   "FB_Z200Conveyor_M211_iDB"(IN_xCycleON := "Z201".ST_xCycleON,
                              IN_xCycleONDel := "Z201".ST_xCycleONDelayed,
                              IN_xFaultsEnabled := "Z201".ST_xFaultsEnabled,
                              IN_xResetAlarms := "Z201".tmOFF_ResetAlarm.OUT_xDone,
                              IN_xAccelation:=FALSE,
                              IN_rgtMotorConfig := #TMP_rgtMotorConfig);
END_REGION

REGION Network 12 (SCL): Outputs Z200
   "ZUPS_Output"();
   "Z201_Output"();
   "Z200_Output"();

   "Output_Z201_Idevice"();
END_REGION
END_ORGANIZATION_BLOCK

// folder: TaskMedium

ORGANIZATION_BLOCK "OBx_TaskMedium"   // OB31, LAD, CyclicInterrupt
{ S7_Optimized_Access := 'TRUE' }
VERSION : 0.1
   VAR_INPUT
      Initial_Call : Bool;   // Initial call of this OB
      Event_Count : Int;   // Events discarded
   END_VAR
   VAR_TEMP
      TMP_iRetVal : Int;
      TMP_xDummy : Bool;
   END_VAR
BEGIN

REGION Network 1: Initialize
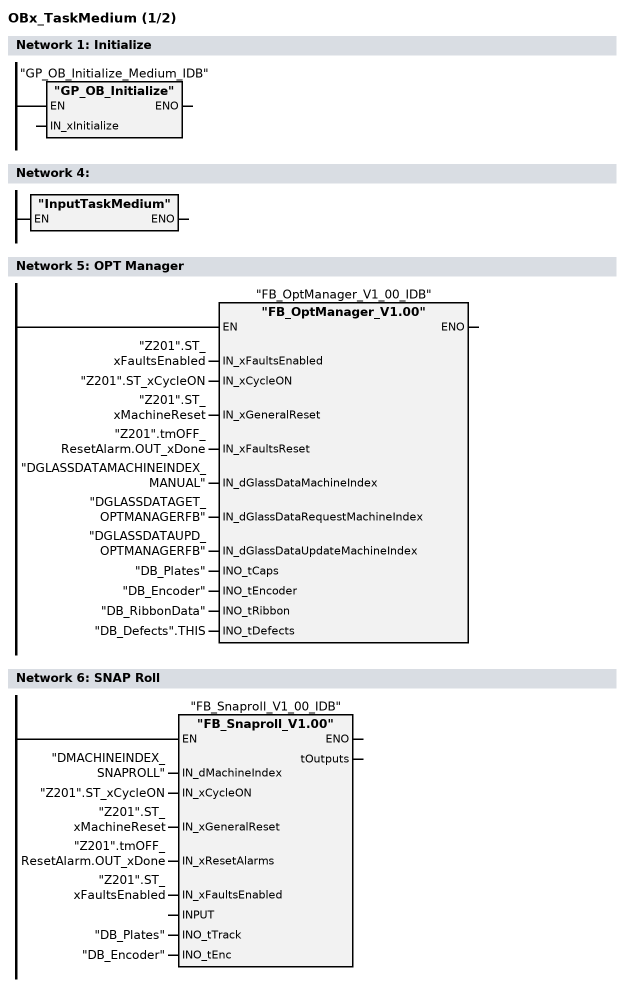
   RUNG wire#powerrail
      "GP_OB_Initialize_Medium_IDB"(IN_xInitialize :=)
   END_RUNG
   // the same network as SCL:
   "GP_OB_Initialize_Medium_IDB"();   // "GP_OB_Initialize"
END_REGION

REGION Network 2: OB Scan
END_REGION

REGION Network 3 (SCL): Message call

   "RP_OB_TaskMediumToOpt"(FALSE);
   "RP_OB_TaskMediumFromOpt"(FALSE);
END_REGION

REGION Network 4
   RUNG wire#powerrail
      "InputTaskMedium"()
   END_RUNG
   // the same network as SCL:
   "InputTaskMedium"();
END_REGION

REGION Network 5: OPT Manager
   RUNG wire#powerrail
      "FB_OptManager_V1_00_IDB"(IN_xFaultsEnabled := "Z201".ST_xFaultsEnabled, IN_xCycleON := "Z201".ST_xCycleON, IN_xGeneralReset := "Z201".ST_xMachineReset, IN_xFaultsReset := "Z201".tmOFF_ResetAlarm.OUT_xDone, IN_dGlassDataMachineIndex := "DGLASSDATAMACHINEINDEX_MANUAL", IN_dGlassDataRequestMachineIndex := "DGLASSDATAGET_OPTMANAGERFB", IN_dGlassDataUpdateMachineIndex := "DGLASSDATAUPD_OPTMANAGERFB", INO_tCaps := "DB_Plates", INO_tEncoder := "DB_Encoder", INO_tRibbon := "DB_RibbonData", INO_tDefects := "DB_Defects".THIS)
   END_RUNG
   // the same network as SCL:
   "FB_OptManager_V1_00_IDB"(IN_xFaultsEnabled := "Z201".ST_xFaultsEnabled,   // "FB_OptManager_V1.00"
                           IN_xCycleON := "Z201".ST_xCycleON,
                           IN_xGeneralReset := "Z201".ST_xMachineReset,
                           IN_xFaultsReset := "Z201".tmOFF_ResetAlarm.OUT_xDone,
                           IN_dGlassDataMachineIndex := "DGLASSDATAMACHINEINDEX_MANUAL",
                           IN_dGlassDataRequestMachineIndex := "DGLASSDATAGET_OPTMANAGERFB",
                           IN_dGlassDataUpdateMachineIndex := "DGLASSDATAUPD_OPTMANAGERFB",
                           INO_tCaps := "DB_Plates",
                           INO_tEncoder := "DB_Encoder",
                           INO_tRibbon := "DB_RibbonData",
                           INO_tDefects := "DB_Defects".THIS);
END_REGION

REGION Network 6: SNAP Roll
   RUNG wire#powerrail
      "FB_Snaproll_V1_00_IDB"(IN_dMachineIndex := "DMACHINEINDEX_SNAPROLL", IN_xCycleON := "Z201".ST_xCycleON, IN_xGeneralReset := "Z201".ST_xMachineReset, IN_xResetAlarms := "Z201".tmOFF_ResetAlarm.OUT_xDone, IN_xFaultsEnabled := "Z201".ST_xFaultsEnabled, INPUT :=, INO_tTrack := "DB_Plates", INO_tEnc := "DB_Encoder", tOutputs =>)
   END_RUNG
   // the same network as SCL:
   "FB_Snaproll_V1_00_IDB"(IN_dMachineIndex := "DMACHINEINDEX_SNAPROLL",   // "FB_Snaproll_V1.00"
                           IN_xCycleON := "Z201".ST_xCycleON,
                           IN_xGeneralReset := "Z201".ST_xMachineReset,
                           IN_xResetAlarms := "Z201".tmOFF_ResetAlarm.OUT_xDone,
                           IN_xFaultsEnabled := "Z201".ST_xFaultsEnabled,
                           INO_tTrack := "DB_Plates",
                           INO_tEnc := "DB_Encoder");
END_REGION

REGION Network 7: Z300
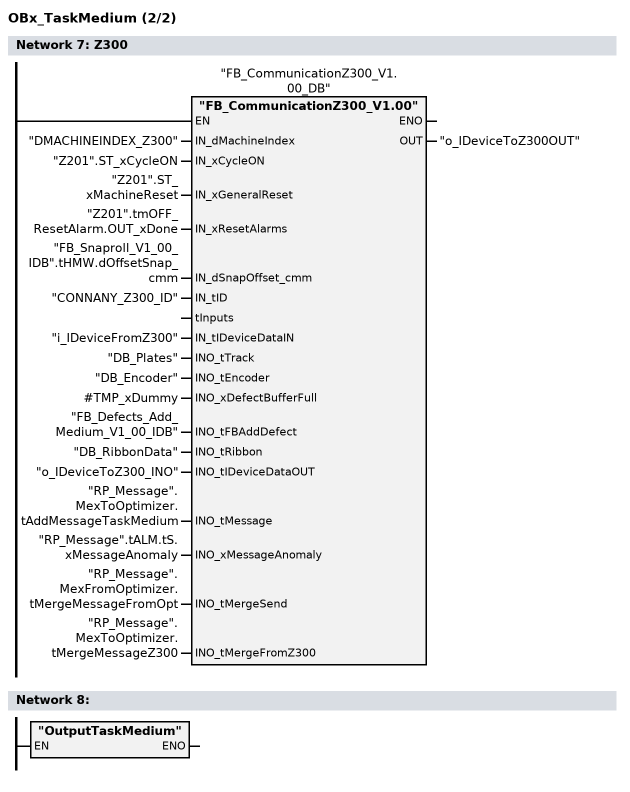
   RUNG wire#powerrail
      "FB_CommunicationZ300_V1.00_DB"(IN_dMachineIndex := "DMACHINEINDEX_Z300", IN_xCycleON := "Z201".ST_xCycleON, IN_xGeneralReset := "Z201".ST_xMachineReset, IN_xResetAlarms := "Z201".tmOFF_ResetAlarm.OUT_xDone, IN_dSnapOffset_cmm := "FB_Snaproll_V1_00_IDB".tHMW.dOffsetSnap_cmm, IN_tID := "CONNANY_Z300_ID", tInputs :=, IN_tIDeviceDataIN := "i_IDeviceFromZ300", INO_tTrack := "DB_Plates", INO_tEncoder := "DB_Encoder", INO_xDefectBufferFull := #TMP_xDummy, INO_tFBAddDefect := "FB_Defects_Add_Medium_V1_00_IDB", INO_tRibbon := "DB_RibbonData", INO_tIDeviceDataOUT := "o_IDeviceToZ300_INO", INO_tMessage := "RP_Message".MexToOptimizer.tAddMessageTaskMedium, INO_xMessageAnomaly := "RP_Message".tALM.tS.xMessageAnomaly, INO_tMergeSend := "RP_Message".MexFromOptimizer.tMergeMessageFromOpt, INO_tMergeFromZ300 := "RP_Message".MexToOptimizer.tMergeMessageZ300, OUT => "o_IDeviceToZ300OUT")
   END_RUNG
   // the same network as SCL:
   "FB_CommunicationZ300_V1.00_DB"(IN_dMachineIndex := "DMACHINEINDEX_Z300",   // "FB_CommunicationZ300_V1.00"
                           IN_xCycleON := "Z201".ST_xCycleON,
                           IN_xGeneralReset := "Z201".ST_xMachineReset,
                           IN_xResetAlarms := "Z201".tmOFF_ResetAlarm.OUT_xDone,
                           IN_dSnapOffset_cmm := "FB_Snaproll_V1_00_IDB".tHMW.dOffsetSnap_cmm,
                           IN_tID := "CONNANY_Z300_ID",
                           IN_tIDeviceDataIN := "i_IDeviceFromZ300",
                           INO_tTrack := "DB_Plates",
                           INO_tEncoder := "DB_Encoder",
                           INO_xDefectBufferFull := #TMP_xDummy,
                           INO_tFBAddDefect := "FB_Defects_Add_Medium_V1_00_IDB",
                           INO_tRibbon := "DB_RibbonData",
                           INO_tIDeviceDataOUT := "o_IDeviceToZ300_INO",
                           INO_tMessage := "RP_Message".MexToOptimizer.tAddMessageTaskMedium,
                           INO_xMessageAnomaly := "RP_Message".tALM.tS.xMessageAnomaly,
                           INO_tMergeSend := "RP_Message".MexFromOptimizer.tMergeMessageFromOpt,
                           INO_tMergeFromZ300 := "RP_Message".MexToOptimizer.tMergeMessageZ300,
                           OUT => "o_IDeviceToZ300OUT");
END_REGION

REGION Network 8
   RUNG wire#powerrail
      "OutputTaskMedium"()
   END_RUNG
   // the same network as SCL:
   "OutputTaskMedium"();
END_REGION
END_ORGANIZATION_BLOCK

// folder: TaskSlow

ORGANIZATION_BLOCK "OBx_TaskSlow"   // OB32, LAD, CyclicInterrupt
{ S7_Optimized_Access := 'TRUE' }
VERSION : 0.1
   VAR_INPUT
      Initial_Call : Bool;   // Initial call of this OB
      Event_Count : Int;   // Events discarded
   END_VAR
   VAR_TEMP
      TMP_xDummy : Bool;
      TMP_iRetVal : Int;
      TMP_rgtMotorConfig : "UDT_MotorConfig";
   END_VAR
BEGIN

REGION Network 1: Initialize
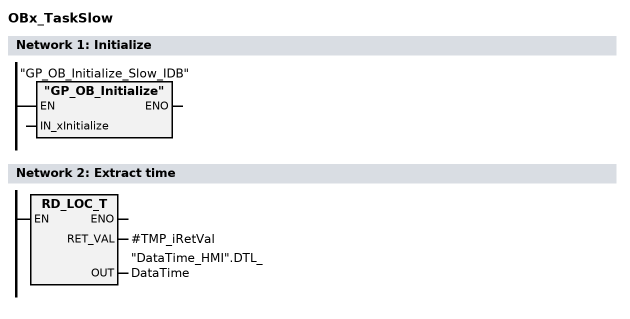
   RUNG wire#powerrail
      "GP_OB_Initialize_Slow_IDB"(IN_xInitialize :=)
   END_RUNG
   // the same network as SCL:
   "GP_OB_Initialize_Slow_IDB"();   // "GP_OB_Initialize"
END_REGION

REGION Network 2: Extract time
   #TMP_iRetVal := RD_LOC_T(OUT => "DataTime_HMI".DTL_DataTime);
END_REGION

REGION Network 3 (SCL)

   "RP_OB_TaskSlowToOpt"(FALSE);

   "RP_OB_TaskSlowFromOpt"(FALSE);

   "InputTaskSlow"();


   "Z200_Logics"();
   "Z200_Faults"();



   "FB_Digitizer_1_V1_00_IDB".IN_tRemoteAddress.ADDR[1] := "IPV4_DIGITIZER_1_IP1";
   "FB_Digitizer_1_V1_00_IDB".IN_tRemoteAddress.ADDR[2] := "IPV4_DIGITIZER_1_IP2";
   "FB_Digitizer_1_V1_00_IDB".IN_tRemoteAddress.ADDR[3] := "IPV4_DIGITIZER_1_IP3";
   "FB_Digitizer_1_V1_00_IDB".IN_tRemoteAddress.ADDR[4] := "IPV4_DIGITIZER_1_IP4";

   "FB_Digitizer_1_V1_00_IDB"(IN_xCycleON:="Z201".ST_xCycleON,
                              IN_xCycleONDel:="Z201".ST_xCycleONDelayed,
                             IN_xGeneralReset:="Z201".ST_xMachineReset,
                             IN_xResetAlarms:="Z201".tmOFF_ResetAlarm.OUT_xDone,
                             IN_xFaultsEnabled:="Z201".ST_xFaultsEnabled,
                             IN_tInterfaceID:="Local~PROFINET_MCC1200",
                             IN_tID:="CONNUOC_DIGITIZER_1",
                             IN_uiRemotePort:="UINT_DIGIITZER_1_PORT",
                             IN_xSimulationActive := "SIMULATION_ACTIVE",  
                             INO_tEnc:="DB_Encoder");

   "FB_Digitizer_2_V1_00_IDB".IN_tRemoteAddress.ADDR[1] := "IPV4_DIGITIZER_2_IP1";
   "FB_Digitizer_2_V1_00_IDB".IN_tRemoteAddress.ADDR[2] := "IPV4_DIGITIZER_2_IP2";
   "FB_Digitizer_2_V1_00_IDB".IN_tRemoteAddress.ADDR[3] := "IPV4_DIGITIZER_2_IP3";
   "FB_Digitizer_2_V1_00_IDB".IN_tRemoteAddress.ADDR[4] := "IPV4_DIGITIZER_2_IP4";

   "FB_Digitizer_2_V1_00_IDB"(IN_xCycleON:="Z201".ST_xCycleON,
                              IN_xCycleONDel:="Z201".ST_xCycleONDelayed,
                             IN_xGeneralReset:="Z201".ST_xMachineReset,
                             IN_xResetAlarms:="Z201".tmOFF_ResetAlarm.OUT_xDone,
                             IN_xFaultsEnabled:="Z201".ST_xFaultsEnabled,
                             IN_tInterfaceID:="Local~PROFINET_MCC1200",
                             IN_tID:="CONNUOC_DIGITIZER_2",
                             IN_uiRemotePort:="UINT_DIGIITZER_2_PORT",
                             IN_xSimulationActive := "SIMULATION_ACTIVE",  
                             INO_tEnc:="DB_Encoder");

   "FB_DigitizerManager_V1_00_IDB"(INO_tDigitizer1:="FB_Digitizer_1_V1_00_IDB",
                                  INO_tDigitizer2:="FB_Digitizer_2_V1_00_IDB",
                                  INO_tEnc:="DB_Encoder",
                                  IN_xCycleON:="Z201".ST_xCycleON,
                                  IN_xCycleONDel:="Z201".ST_xCycleONDelayed,
                                  IN_xGeneralReset:="Z201".ST_xMachineReset,
                                  IN_xResetAlarms:="Z201".tmOFF_ResetAlarm.OUT_xDone,
                                  IN_xFaultsEnabled:="Z201".ST_xFaultsEnabled);


   "FB_YCuts1_V1_00_IDB"(IN_dMachineIndex:="DMACHINEINDEX_YCUT1",
                        IN_dYCUTID:=0,
                        IN_dTrackNewCapIndex:="DINDEXNEWCAPAVAILABLE_YCUT1",
                        IN_xCycleON:="Z201".ST_xCycleON,
                        IN_xGeneralReset:="Z201".ST_xMachineReset,
                        IN_xResetAlarms:="Z201".tmOFF_ResetAlarm.OUT_xDone,
                        IN_xFaultsEnabled:="Z201".ST_xFaultsEnabled,
                        IN_tID:="CONNANY_YCUT1_ID",

                        IN_dGlassBreakMachineIndex := "DGLASSBREAKGET_YCUT1",
                        INO_tTrack:="DB_Plates",
                        INO_tEnc:="DB_Encoder",
                        INO_tRibbon := "DB_RibbonData",
                        IN_xSimulationActive:= "SIMULATION_ACTIVE");

   "FB_YCuts2_V1_00_IDB"(IN_dMachineIndex:="DMACHINEINDEX_YCUT2",
                        IN_dYCUTID:=1,
                        IN_dTrackNewCapIndex:="DINDEXNEWCAPAVAILABLE_YCUT2",
                        IN_xCycleON:="Z201".ST_xCycleON,
                        IN_xGeneralReset:="Z201".ST_xMachineReset,
                        IN_xResetAlarms:="Z201".tmOFF_ResetAlarm.OUT_xDone,
                        IN_xFaultsEnabled:="Z201".ST_xFaultsEnabled,
                        IN_tID:="CONNANY_YCUT2_ID",
                        IN_dGlassBreakMachineIndex := "DGLASSBREAKGET_YCUT2",   
                        INO_tTrack:="DB_Plates",
                        INO_tEnc:="DB_Encoder",
                        INO_tRibbon := "DB_RibbonData",
                        IN_xSimulationActive:= "SIMULATION_ACTIVE");



   "FB_CrossCuts_1_V1_00_IDB"(IN_dMachineIndex:="DMACHINEINDEX_XCUT1",
                              IN_dGlassSearchMachineIndex_Q0:="DGLASSSEARCHMACHINEINDEX_XCUT1_Q0",
                              IN_dGlassSearchMachineIndex_Q1:="DGLASSSEARCHMACHINEINDEX_XCUT1_Q1",
                              IN_dGlassSearchMachineIndex_Q2:="DGLASSSEARCHMACHINEINDEX_XCUT1_Q2",
                              IN_dGlassSearchMachineIndex_Q3:="DGLASSSEARCHMACHINEINDEX_XCUT1_Q3",
                              IN_dXCutIndex := 0,
                              IN_xCycleON:="Z201".ST_xCycleON,
                              IN_xGeneralReset:="Z201".ST_xMachineReset,
                              IN_xResetAlarms:="Z201".tmOFF_ResetAlarm.OUT_xDone,
                              IN_xFaultsEnabled:="Z201".ST_xFaultsEnabled,
                              IN_xSimulationActive:= "SIMULATION_ACTIVE",
                              INO_tTrack:="DB_Plates",
                              INO_tOBInit := "GP_OB_Initialize_Slow_IDB",
                              INO_tRibbon := "DB_RibbonData",
                              INO_tEnc:="DB_Encoder",
                              INO_tXCutOpt:= "FB_CrossCut_Opt_V1_00_IDB" ,
                              IN_dGlassBreakMachineIndex := "DGLASSBREAKGET_XCUT1",
                              IN_xMBDone:="DB_XCut1_MBClientInstance".DONE,
                              IN_xMBError:="DB_XCut1_MBClientInstance".ERROR);

   "FB_CrossCuts_2_V1_00_IDB"(IN_dMachineIndex:="DMACHINEINDEX_XCUT2",
                              IN_dGlassSearchMachineIndex_Q0:="DGLASSSEARCHMACHINEINDEX_XCUT2_Q0",
                              IN_dGlassSearchMachineIndex_Q1:="DGLASSSEARCHMACHINEINDEX_XCUT2_Q1",
                              IN_dGlassSearchMachineIndex_Q2:="DGLASSSEARCHMACHINEINDEX_XCUT2_Q2",
                              IN_dGlassSearchMachineIndex_Q3:="DGLASSSEARCHMACHINEINDEX_XCUT2_Q3",
                              IN_dXCutIndex := 1,
                              IN_xCycleON:="Z201".ST_xCycleON,
                              IN_xGeneralReset:="Z201".ST_xMachineReset,
                              IN_xResetAlarms:="Z201".tmOFF_ResetAlarm.OUT_xDone,
                              IN_xFaultsEnabled:="Z201".ST_xFaultsEnabled,
                              IN_xSimulationActive:= "SIMULATION_ACTIVE",
                              INO_tTrack:="DB_Plates",
                              INO_tOBInit := "GP_OB_Initialize_Slow_IDB",
                              INO_tRibbon := "DB_RibbonData",
                              INO_tEnc:="DB_Encoder",
                              INO_tXCutOpt:= "FB_CrossCut_Opt_V1_00_IDB",
                              IN_dGlassBreakMachineIndex := "DGLASSBREAKGET_XCUT2",
                              IN_xMBDone:="DB_XCut2_MBClientInstance".DONE,
                              IN_xMBError:="DB_XCut2_MBClientInstance".ERROR);

   "FB_CrossCuts_3_V1_00_IDB"(IN_dMachineIndex := "DMACHINEINDEX_XCUT3",
                              IN_dGlassSearchMachineIndex_Q0 := "DGLASSSEARCHMACHINEINDEX_XCUT3_Q0",
                              IN_dGlassSearchMachineIndex_Q1 := "DGLASSSEARCHMACHINEINDEX_XCUT3_Q1",
                              IN_dGlassSearchMachineIndex_Q2 := "DGLASSSEARCHMACHINEINDEX_XCUT3_Q2",
                              IN_dGlassSearchMachineIndex_Q3 := "DGLASSSEARCHMACHINEINDEX_XCUT3_Q3",
                              IN_dXCutIndex := 1,
                              IN_xCycleON := "Z201".ST_xCycleON,
                              IN_xGeneralReset := "Z201".ST_xMachineReset,
                              IN_xResetAlarms := "Z201".tmOFF_ResetAlarm.OUT_xDone,
                              IN_xFaultsEnabled := "Z201".ST_xFaultsEnabled,
                              IN_xSimulationActive := "SIMULATION_ACTIVE",
                              INO_tTrack := "DB_Plates",
                              INO_tOBInit := "GP_OB_Initialize_Slow_IDB",
                              INO_tRibbon := "DB_RibbonData",
                              INO_tEnc := "DB_Encoder",
                              INO_tXCutOpt := "FB_CrossCut_Opt_V1_00_IDB",
                              IN_dGlassBreakMachineIndex := "DGLASSBREAKGET_XCUT3",
                              IN_xMBDone := "DB_XCut3_MBClientInstance".DONE,
                              IN_xMBError := "DB_XCut3_MBClientInstance".ERROR);


   "FB_Markers_V1.00_IDB"(IN_xStandardFBCall:=TRUE,
                         IN_xCycleON:="Z201".ST_xCycleON,
                         IN_xGeneralReset:="Z201".ST_xMachineReset,
                         IN_xResetAlarms:="Z201".tmOFF_ResetAlarm.OUT_xDone,
                         IN_xFaultsEnabled:="Z201".ST_xFaultsEnabled,
                         IN_tID:="CONNANY_MARKER_ID",
                         IN_dGlassBreakMachineIndex:="DGLASSBREAKGET_MARKER",
                         INO_tEnc:="DB_Encoder",
                         INO_tRibbon:="DB_RibbonData");



   "FB_BD_BreakPH_V1_00_IDB"(IN_xCycleON:="ZUPS".ST_xCycleON,
                             IN_xCycleONDel:="ZUPS".ST_xCycleONDelayed,
                             IN_xGeneralReset:="Z201".ST_xMachineReset,
                          IN_xResetAlarms:="Z201".tmOFF_ResetAlarm.OUT_xDone,
                          IN_xFaultsEnabled:="ZUPS".ST_xFaultsEnabled,
                          IN_dNumUsedPhoto:=10,
                          IN_dIndexBreakMachine:="DGLASSBREAKMACHINEINDEX_M202",
                          INO_tEncoder:="DB_Encoder",
                          INO_tFBAddDefect := "FB_Defects_Add_Slow_V1_00_IDB",
                          INO_tRibbon:="DB_RibbonData");


   "FB_BD_DigitizerPH_V1_00_IDB".tHMW.dMinBreakSize_cmm := 2000;
   "FB_BD_DigitizerPH_V1_00_IDB".tHMW.dDistanceSnaproll_cmm := 1121200;
   "FB_BD_DigitizerPH_V1_00_IDB".tHMR.dDistanceSnaproll_cmm := 1121200;

   IF "FB_Digitizer_1_V1_00_IDB".tHMW.xGlassSensorEnabled AND NOT "FB_Digitizer_1_V1_00_IDB".tHMR.xManComEn THEN
       "FB_BD_DigitizerPH_V1_00_IDB".tHMR.rgdPhotoAbilitation[0] := 3;
   ELSE
       "FB_BD_DigitizerPH_V1_00_IDB".tHMR.rgdPhotoAbilitation[0] := 1;
   END_IF;

   IF "FB_Digitizer_2_V1_00_IDB".tHMW.xGlassSensorEnabled AND NOT "FB_Digitizer_2_V1_00_IDB".tHMR.xManComEn THEN
       "FB_BD_DigitizerPH_V1_00_IDB".tHMR.rgdPhotoAbilitation[1] := 3;
   ELSE
       "FB_BD_DigitizerPH_V1_00_IDB".tHMR.rgdPhotoAbilitation[1] := 1;
   END_IF;


   "FB_BD_DigitizerPH_V1_00_IDB"(IN_xCycleON := "Z201".ST_xCycleON,
                               IN_xCycleONDel := "Z201".ST_xCycleONDelayed,
                          IN_xGeneralReset := "Z201".ST_xMachineReset,
                          IN_xResetAlarms := "Z201".tmOFF_ResetAlarm.OUT_xDone,
                          IN_xFaultsEnabled := "Z201".ST_xFaultsEnabled,
                          IN_dNumUsedPhoto := 2,
                          IN_dIndexBreakMachine := "DGLASSBREAKMACHINEINDEX_M216",
                          INO_tEncoder := "DB_Encoder",
                          INO_tFBAddDefect := "FB_Defects_Add_Slow_V1_00_IDB",
                          INO_tRibbon := "DB_RibbonData");

   "FB_ColdBackupManager_V1_00_DB"(IN_xGeneralReset:="Z201".ST_xMachineReset,
                                   IN_xResetAlarms:="Z201".tmOFF_ResetAlarm.OUT_xDone,
                                   IN_tHWInterface:="Local~PROFINET_MCC1200~Port_2",
                                   IN_xThisPLCActive:="Z201".ST_xThisPlcActive);

   "ExChangeParTxRx_Logic"(IN_tConfDataBackup := "FB_ColdBackupManager_V1_00_DB".IN_tConfDataBackup,
                           IN_tConfDataMaster := "FB_ColdBackupManager_V1_00_DB".IN_tConfDataMaster);

   "FB_Oil_V1_00_IDB"(IN_xCycleON:="Z201".ST_xCycleON,
                      IN_xCycleONDel:="Z201".ST_xCycleONDelayed,
                      IN_xGeneralReset:="Z201".ST_xMachineReset,
                      IN_xResetAlarms:="Z201".tmOFF_ResetAlarm.OUT_xDone,
                      IN_xFaultsEnabled:="Z201".ST_xFaultsEnabled,
                      INO_tOBInitialize:="GP_OB_Initialize_Slow_IDB");

   "FB_ManInsp_V1_00_IDB"(IN_xCycleON:="Z201".ST_xCycleON,
                          IN_dNumButtonDefect := 12,
                          IN_dNumQltDefect := 4,
                          INO_tEncoder := "DB_Encoder",
                          INO_tFBAddDefect := "FB_Defects_Add_Slow_V1_00_IDB",
                          INO_xDefectBufferFull := #TMP_xDummy,
                          IN_xCycleONDel:="Z201".ST_xCycleONDelayed,
                          IN_xGeneralReset:="Z201".ST_xMachineReset,
                          IN_xResetAlarms:="Z201".tmOFF_ResetAlarm.OUT_xDone,
                          IN_xFaultsEnabled:="Z201".ST_xFaultsEnabled,
                          IN_dGlassBreakMachineIndex :="DGLASSBREAKMACHINEINDEX_M212",
                          INO_tRibbon := "DB_RibbonData",
                          INO_tOBInitialize:="GP_OB_Initialize_Slow_IDB");

   "FB_WanderCamera_V1_00_IDB".IN_tRemoteAddress.ADDR[1] := "IPV4_WANDER_IP1";
   "FB_WanderCamera_V1_00_IDB".IN_tRemoteAddress.ADDR[2] := "IPV4_WANDER_IP2";
   "FB_WanderCamera_V1_00_IDB".IN_tRemoteAddress.ADDR[3] := "IPV4_WANDER_IP3";
   "FB_WanderCamera_V1_00_IDB".IN_tRemoteAddress.ADDR[4] := "IPV4_WANDER_IP4";

   "FB_WanderCamera_V1_00_IDB"(IN_xCycleON := "Z201".ST_xCycleON,
                               IN_xCycleONDel := "Z201".ST_xCycleONDelayed,
                               IN_xGeneralReset := "Z201".ST_xMachineReset,
                               IN_xResetAlarms := "Z201".tmOFF_ResetAlarm.OUT_xDone,
                               IN_xFaultsEnabled := "Z201".ST_xFaultsEnabled,
                               IN_dGlassBreakMachineIndex := "DMACHINEINDEX_GETGLASSBREAK_WANDER",
                               IN_dGlassDataMachineIndex := "DGLASSDATAMACHINEINDEX_CAMERA",
                               IN_tInterfaceID := "Local~PROFINET_MCC1200~Port_2",
                               IN_tID := "CONNUOC_WANDER",
                               IN_uiRemotePort := "UINT_WANDER_PORT",
                               INO_tRibbon := "DB_RibbonData",
                               INO_tTrack := "DB_Plates");

   "FB_ISRA5D_IDB"(IN_xCycleON := "Z201".ST_xCycleON,
                   IN_xCycleONDel := "Z201".ST_xCycleONDelayed,
                   IN_xGeneralReset := "Z201".ST_xMachineReset,
                   IN_xResetAlarms := "Z201".tmOFF_ResetAlarm.OUT_xDone,
                   IN_xFaultsEnabled := "Z201".ST_xFaultsEnabled,
                   IN_tID := "CONNUOC_ISRA5D",
                   IN_tInterfaceID := "Local~PCNETWORK_MCC1200",
                   IN_uiLocalPort := "UINT_ISRA5D_PORT",
                   IN_dGlassBreakIndexGet := "DGLASSBREAKGET_ISRA5DFB",
                   IN_dGlassDataMachineIndex :="DGLASSDATAMACHINEINDEX_SCANNER" ,
                   IN_dGlassDataUpdateMachineIndex := "DGLASSDATAUPD_ISRA5DFB",
                   IN_xSimulationActive := FALSE,
                   INO_OB_Init := "GP_OB_Initialize_Slow_IDB",
                   INO_tCaps := "DB_Plates",
                   INO_tEncoder := "DB_Encoder",
                   INO_tFBAddDefect := "FB_Defects_Add_Slow_V1_00_IDB",
                   INO_tOptManager := "FB_OptManager_V1_00_IDB",
                   INO_tRibbon := "DB_RibbonData",
                   INO_xDefectBufferFull := #TMP_xDummy);





   //"FB_DropConveyor_IDB"(IN_xCycleON := "ZUPS".ST_xCycleON,
                        // IN_xCycleONDel := "ZUPS".ST_xCycleONDelayed,
                       //  IN_xResetAlarms := "Z201".tmOFF_ResetAlarm.OUT_xDone,
                      //   IN_xFaultsEnabled := "ZUPS".ST_xFaultsEnabled,
                      //   IN_xManualMode := "FB_Z200Conveyor_M203_IDB".tHMR.xManualCommandEnabled,
                     //    IN_dActualLehrSpeed_mm_min := "FB_LehrSpeed_IDB".tHMR.dActualSpeedValue_mm_min,
                    //     IN_dGlassBreakMachineIndex := "DGLASSBREAKMACHINEINDEX_M204",
                     //    IN_xSimulationActive := "SIMULATION_ACTIVE",
                     //    INO_tRibbon := "DB_RibbonData");

   //"FB_BreakerM205_V1.00_IDB"(IN_xCycleON := "ZUPS".ST_xCycleON,
              //                IN_xCycleONDel := "ZUPS".ST_xCycleONDelayed,
                        //      IN_xGeneralReset := "Z201".ST_xMachineReset,
                        //      IN_xResetAlarms := "Z201".tmOFF_ResetAlarm.OUT_xDone,
                         //     IN_xFaultsEnabled := "ZUPS".ST_xFaultsEnabled,
                        //      IN_xDropConveyorDown := "FB_DropConveyor_IDB".tHMR.xDownPosition,
                        //      INO_tOBInitialize := "GP_OB_Initialize_Slow_IDB");


   "Z200_SpeedLehr"();
END_REGION

REGION Network 4 (SCL): Outputs


   "OutputTaskSlow"();
END_REGION
END_ORGANIZATION_BLOCK

// folder: TaskStartup

ORGANIZATION_BLOCK "Startup"   // OB100, LAD, Startup
TITLE = "Complete Restart"
{ S7_Optimized_Access := 'TRUE' }
VERSION : 0.1
   VAR_INPUT
      LostRetentive : Bool;   // True if retentive data are lost
      LostRTC : Bool;   // True if date and time are lost
   END_VAR
BEGIN

REGION Network 1 (SCL): Initialization
   //Initialize all FB
   "DB_Z201_HMI".tHMW.xGeneralReset := TRUE;
   "Z201".ST_xMachineReset:= TRUE;
   "GP_OB_Initialize_Fast_IDB".IN_xInitialize := TRUE;
   "GP_OB_Initialize_Medium_IDB".IN_xInitialize := TRUE;
   "GP_OB_Initialize_Slow_IDB".IN_xInitialize := TRUE;
   "GP_OB_Initialize_Fast_IDB".IN_xInitialize := TRUE;

   //Inizializa all reports
   "RP_OB_TaskFastFromOpt"(TRUE);
   "RP_OB_TaskFastToOpt"(TRUE);
   "RP_OB_TaskMainFromOpt"(TRUE);
   "RP_OB_TaskMainToOpt"(TRUE);
   "RP_OB_TaskMediumFromOpt"(TRUE);
   "RP_OB_TaskMediumToOpt"(TRUE);
   "RP_OB_TaskSlowFromOpt"(TRUE);
   "RP_OB_TaskSlowToOpt"(TRUE);

   //Compile data for redundancy manager
   "FB_ColdBackupManager_V1_00_DB".IN_tConfDataMaster.Header.SubfieldCount := 1;
   "FB_ColdBackupManager_V1_00_DB".IN_tConfDataMaster.IPData.Mode := 1;
   "FB_ColdBackupManager_V1_00_DB".IN_tConfDataMaster.IPData.InterfaceAddress.ADDR[1] := 192;
   "FB_ColdBackupManager_V1_00_DB".IN_tConfDataMaster.IPData.InterfaceAddress.ADDR[2] := 168;
   "FB_ColdBackupManager_V1_00_DB".IN_tConfDataMaster.IPData.InterfaceAddress.ADDR[3] := 130;
   "FB_ColdBackupManager_V1_00_DB".IN_tConfDataMaster.IPData.InterfaceAddress.ADDR[4] := 5;
   "FB_ColdBackupManager_V1_00_DB".IN_tConfDataMaster.IPData.SubnetMask.ADDR[1] := 255;
   "FB_ColdBackupManager_V1_00_DB".IN_tConfDataMaster.IPData.SubnetMask.ADDR[2] := 255;
   "FB_ColdBackupManager_V1_00_DB".IN_tConfDataMaster.IPData.SubnetMask.ADDR[3] := 255;
   "FB_ColdBackupManager_V1_00_DB".IN_tConfDataMaster.IPData.SubnetMask.ADDR[4] := 0;


   "FB_ColdBackupManager_V1_00_DB".IN_tConfDataBackup.Header.SubfieldCount := 1;
   "FB_ColdBackupManager_V1_00_DB".IN_tConfDataBackup.IPData.Mode := 1;
   "FB_ColdBackupManager_V1_00_DB".IN_tConfDataBackup.IPData.InterfaceAddress.ADDR[1] := 192;
   "FB_ColdBackupManager_V1_00_DB".IN_tConfDataBackup.IPData.InterfaceAddress.ADDR[2] := 168;
   "FB_ColdBackupManager_V1_00_DB".IN_tConfDataBackup.IPData.InterfaceAddress.ADDR[3] := 130;
   "FB_ColdBackupManager_V1_00_DB".IN_tConfDataBackup.IPData.InterfaceAddress.ADDR[4] := 6;
   "FB_ColdBackupManager_V1_00_DB".IN_tConfDataBackup.IPData.SubnetMask.ADDR[1] := 255;
   "FB_ColdBackupManager_V1_00_DB".IN_tConfDataBackup.IPData.SubnetMask.ADDR[2] := 255;
   "FB_ColdBackupManager_V1_00_DB".IN_tConfDataBackup.IPData.SubnetMask.ADDR[3] := 255;
   "FB_ColdBackupManager_V1_00_DB".IN_tConfDataBackup.IPData.SubnetMask.ADDR[4] := 0;

   //Initialize tracking plate data
   "DB_Plates".tNewCapToInsert := "DB_Plates".tEmptyCap;

   "DB_Plates".tNewCapToInsert.dLength_cmm := 200000;
   "DB_Plates".tNewCapToInsert.dWidth_cmm := 321000;
   "DB_Plates".tNewCapToInsert.dThick_cmm := 500;
   "DB_Plates".tNewCapToInsert.dNumLites := 1;
   "DB_Plates".tNewCapToInsert.rgtLites[0].dWidth_cmm := 321000;

   //Initialize Ribbon data buffer
   "DB_RibbonData".dActualNumberGlassBreakMachine := 3;
   "DB_RibbonData".dActualNumberGlassDataMachine := 3;

   "DB_RibbonData".rgtGlassBreak[0].dDistSnapRoll_cmm := "FB_BD_BreakPH_V1_00_IDB".tHMR.dDistanceSnaproll_cmm;
   "DB_RibbonData".rgtGlassBreak[1].dDistSnapRoll_cmm := "FB_BD_DigitizerPH_V1_00_IDB".tHMR.dDistanceSnaproll_cmm;
END_REGION
END_ORGANIZATION_BLOCK

// ===== PLC "2B160AP"  CPU 1512SP-1 PN =====

VAR_GLOBAL   // PLC tag table "Tabella delle variabili standard"
   "AlwaysFALSE" AT %M0.3 : Bool;
   "AlwaysOFF_Debug" AT %M10.0 : Bool;
   "AlwaysTRUE" AT %M0.2 : Bool;
   "cigliu" AT %M1.0 : Bool;
   "DiagStatusUpdate" AT %M0.1 : Bool;
   "FirstScan" AT %M0.0 : Bool;
   "i.1B160AP1.1B11QF1/2.AnomalyPowerSupplies230V" AT %E0.2 : Bool;
   "i.1B160AP1.1B18-2L+.PowerSupplyInputControlCabinetON" AT %E0.0 : Bool;
   "i.1B160AP1.1B18-3L+.InputInstallationPowerSupplyON" AT %E0.1 : Bool;
   "i.1B160AP1.1B18QF2.PowerSupply24VLogic" AT %E0.3 : Bool;
   "i.1B160AP1.1B18QF3.PowerSupply24VLogic" AT %E0.4 : Bool;
   "i.1B160AP1.1B20QF2.PowerSupply24VLogic" AT %E0.5 : Bool;
   "i.1B160AP1.1B20QF3.PowerSupply24VLogic" AT %I0.6 : Bool;
   "i.1B160AP1.1B122KE1.MainEmergencyON" AT %E1.1 : Bool;
   "i.1B160AP1.1B41QF1.ProtectionPowerSupply36V_Motor_1-4" AT %I1.4 : Bool;
   "i.1B160AP1.1B41QF2.ProtectionPowerSupplyMotorsYcut_1-4" AT %I1.5 : Bool;
   "i.1B160AP1.1B42QF1.ProtectionPowerSupply36V_Motor_5-8" AT %I1.6 : Bool;
   "i.1B160AP1.1B42QF2.ProtectionPowerSupplyMotorsYcut_5-8" AT %I1.7 : Bool;
   "i.1B160AP1.1B51QM1.ProtectionCarriageTranslation" AT %E2.0 : Bool;
   "i.1B160AP1.1B52QM1.ProtectionCarriageTranslation" AT %E2.1 : Bool;
   "i.1B160AP1.1B53QM1.ProtectionCarriageTranslation" AT %E2.2 : Bool;
   "i.1B160AP1.1B54QM1.ProtectionCarriageTranslation" AT %E2.3 : Bool;
   "i.1B160AP1.1B55QM1.ProtectionCarriageTranslation" AT %I2.4 : Bool;
   "i.1B160AP1.1B56QM1.ProtectionCarriageTranslation" AT %I2.5 : Bool;
   "i.1B160AP1.1B57QM1.ProtectionCarriageTranslation" AT %I2.6 : Bool;
   "i.1B160AP1.1B58QM1.ProtectionCarriageTranslation" AT %I2.7 : Bool;
   "i.1B160AP1.M217B1SB1.LocalEmergency" AT %I3.1 : Bool;
   "i.1B160AP1.M217B1SB2.LocalEmergency" AT %I3.2 : Bool;
   "i.1B160AP1.M217B1SB3_SB4.HeadsUpIstantaneous" AT %I3.0 : Bool;
   "i.1B406AP1.1B406SB4.HeadsUpIstantaneous" AT %E106.3 : Bool;
   "i.1B160AP1.CaptureValue" AT %ID34 : DWord;
   "i.1B160AP1.CounterActualValue" AT %ID30 : DWord;
   "i.1B160AP1.CounterCardStatus" AT %ED42 : DWord;
   "i.1B160AP1.Event_Capture" AT %I45.6 : Bool;
   "i.1B160AP1.FrequencyActualValue" AT %ID38 : Real;
   "i.1B160AP1.Res_Event_Ack" AT %I43.1 : Bool;
   "i.1B411AP1.1B411SA1.Head1.CuttingPressure-" AT %E112.2 : Bool;
   "i.1B411AP1.1B411SA1.Head1.CuttingPressure+" AT %E111.2 : Bool;
   "i.1B411AP1.1B411SA2.Head1.ProductionON" AT %E112.4 : Bool;
   "i.1B411AP1.1B411SQ1.Head1.CarriageHeadWorkPosition" AT %E111.3 : Bool;
   "i.1B412AP1.1B412SA1.Head2.CuttingPressure-" AT %E122.2 : Bool;
   "i.1B412AP1.1B412SA1.Head2.CuttingPressure+" AT %E121.2 : Bool;
   "i.1B412AP1.1B412SA2.Head2.ProductionON" AT %E122.4 : Bool;
   "i.1B412AP1.1B412SQ1.Head2.CarriageHeadWorkPosition" AT %E121.3 : Bool;
   "i.1B413AP1.1B413SA1.Head3.CuttingPressure-" AT %E132.2 : Bool;
   "i.1B413AP1.1B413SA1.Head3.CuttingPressure+" AT %E131.2 : Bool;
   "i.1B413AP1.1B413SA2.Head3.ProductionON" AT %E132.4 : Bool;
   "i.1B413AP1.1B413SQ1.Head3.CarriageHeadWorkPosition" AT %E131.3 : Bool;
   "i.1B414AP1.1B414SA1.Head4.CuttingPressure-" AT %E142.2 : Bool;
   "i.1B414AP1.1B414SA1.Head4.CuttingPressure+" AT %E141.2 : Bool;
   "i.1B414AP1.1B414SA2.Head4.ProductionON" AT %E142.4 : Bool;
   "i.1B414AP1.1B414SQ1.Head4.CarriageHeadWorkPosition" AT %E141.3 : Bool;
   "i.1B415AP1.1B415SA1.Head5.CuttingPressure-" AT %I152.2 : Bool;
   "i.1B415AP1.1B415SA1.Head5.CuttingPressure+" AT %I151.2 : Bool;
   "i.1B415AP1.1B415SA2.Head5.ProductionON" AT %I152.4 : Bool;
   "i.1B415AP1.1B415SQ1.Head5.CarriageHeadWorkPosition" AT %I151.3 : Bool;
   "i.1B416AP1.1B416SA1.Head6.CuttingPressure-" AT %I162.2 : Bool;
   "i.1B416AP1.1B416SA1.Head6.CuttingPressure+" AT %I161.2 : Bool;
   "i.1B416AP1.1B416SA2.Head6.ProductionON" AT %I162.4 : Bool;
   "i.1B416AP1.1B416SQ1.Head6.CarriageHeadWorkPosition" AT %I161.3 : Bool;
   "i.1B417AP1.1B417SA1.Head7.CuttingPressure-" AT %I172.2 : Bool;
   "i.1B417AP1.1B417SA1.Head7.CuttingPressure+" AT %I171.2 : Bool;
   "i.1B417AP1.1B417SA2.Head7.ProductionON" AT %I172.4 : Bool;
   "i.1B417AP1.1B417SQ1.Head7.CarriageHeadWorkPosition" AT %I171.3 : Bool;
   "i.1B418AP1.1B418SA1.Head8.CuttingPressure-" AT %I182.2 : Bool;
   "i.1B418AP1.1B418SA1.Head8.CuttingPressure+" AT %I181.2 : Bool;
   "i.1B418AP1.1B418SA2.Head8.ProductionON" AT %I182.4 : Bool;
   "i.1B418AP1.1B418SQ1.Head8.CarriageHeadWorkPosition" AT %I181.3 : Bool;
   "i.IDeviceCPU0" AT %I250.0 : "UDT_CM_IDEV_FromMainLine";
   "o.1B160AP1.1B251HL1.AreaFailure" AT %A0.0 : Bool;
   "o.1B160AP1.1B251KA1.ResetLocalEmergency" AT %A0.2 : Bool;
   "o.1B160AP1.EnableCard1" AT %A2.0 : Bool;
   "o.1B160AP1.EnableCard2" AT %A2.1 : Bool;
   "o.1B160AP1.EnableCard3" AT %A2.2 : Bool;
   "o.1B160AP1.EnableCard4" AT %A2.3 : Bool;
   "o.1B160AP1.EnableCard5" AT %Q2.4 : Bool;
   "o.1B160AP1.EnableCard6" AT %Q2.5 : Bool;
   "o.1B160AP1.EnableCard7" AT %Q2.6 : Bool;
   "o.1B160AP1.EnableCard8" AT %Q2.7 : Bool;
   "o.1B160AP1.M217B1HL3.MachineReady" AT %Q0.4 : Bool;
   "o.1B160AP1.M217B1HL4.MachineInOrder" AT %Q0.5 : Bool;
   "o.1B160AP1.M217B1HL5.MachineToMaintenance" AT %Q0.6 : Bool;
   "o.1B160AP1.M217B1HL6.MachineOutOfOrder" AT %Q0.7 : Bool;
   "o.1B160AP1.M217CutPressureHead1" AT %AW50 : Int;
   "o.1B160AP1.M217CutPressureHead2" AT %AW52 : Int;
   "o.1B160AP1.M217CutPressureHead3" AT %AW54 : Int;
   "o.1B160AP1.M217CutPressureHead4" AT %QW56 : Int;
   "o.1B160AP1.M217CutPressureHead5" AT %QW58 : Int;
   "o.1B160AP1.M217CutPressureHead6" AT %QW60 : Int;
   "o.1B160AP1.M217CutPressureHead7" AT %QW62 : Int;
   "o.1B160AP1.M217CutPressureHead8" AT %QW64 : Int;
   "o.1B160AP1.CounterCardStatus" AT %AD38 : DWord;
   "o.1B160AP1.Enable_Measure" AT %Q39.7 : Bool;
   "o.1B160AP1.Open_SW_Gate" AT %Q39.0 : Bool;
   "o.1B160AP1.Res_Event" AT %Q40.1 : Bool;
   "o.1B411AP1.1B411SA2.Head1.ProductionON" AT %A111.4 : Bool;
   "o.1B411AP1.1B411YV1.Head1.CuttingHeadGlassApproach" AT %A111.1 : Bool;
   "o.1B411AP1.1B411YV2.Head1.CuttingLubrication" AT %A111.0 : Bool;
   "o.1B412AP1.1B412SA2.Head2.ProductionON" AT %A121.4 : Bool;
   "o.1B412AP1.1B412YV1.Head2.CuttingHeadGlassApproach" AT %A121.1 : Bool;
   "o.1B412AP1.1B412YV2.Head2.CuttingLubrication" AT %A121.0 : Bool;
   "o.1B413AP1.1B413SA2.Head3.ProductionON" AT %A131.4 : Bool;
   "o.1B413AP1.1B413YV1.Head3.CuttingHeadGlassApproach" AT %A131.1 : Bool;
   "o.1B413AP1.1B413YV2.Head3.CuttingLubrication" AT %A131.0 : Bool;
   "o.1B414AP1.1B414SA2.Head4.ProductionON" AT %A141.4 : Bool;
   "o.1B414AP1.1B414YV1.Head4.CuttingHeadGlassApproach" AT %A141.1 : Bool;
   "o.1B414AP1.1B414YV2.Head4.CuttingLubrication" AT %A141.0 : Bool;
   "o.1B415AP1.1B415SA2.Head5.ProductionON" AT %Q151.4 : Bool;
   "o.1B415AP1.1B415YV1.Head5.CuttingHeadGlassApproach" AT %Q151.1 : Bool;
   "o.1B415AP1.1B415YV2.Head5.CuttingLubrication" AT %Q151.0 : Bool;
   "o.1B416AP1.1B416SA2.Head6.ProductionON" AT %Q161.4 : Bool;
   "o.1B416AP1.1B416YV1.Head6.CuttingHeadGlassApproach" AT %Q161.1 : Bool;
   "o.1B416AP1.1B416YV2.Head6.CuttingLubrication" AT %Q161.0 : Bool;
   "o.1B417AP1.1B417SA2.Head7.ProductionON" AT %Q171.4 : Bool;
   "o.1B417AP1.1B417YV1.Head7.CuttingHeadGlassApproach" AT %Q171.1 : Bool;
   "o.1B417AP1.1B417YV2.Head7.CuttingLubrication" AT %Q171.0 : Bool;
   "o.1B418AP1.1B418SA2.Head8.ProductionON" AT %Q181.4 : Bool;
   "o.1B418AP1.1B418YV1.Head8.CuttingHeadGlassApproach" AT %Q181.1 : Bool;
   "o.1B418AP1.1B418YV2.Head8.CuttingLubrication" AT %Q181.0 : Bool;
   "o.IDeviceCPU0" AT %Q250.0 : "UDT_CM_IDEV_ToMainLine";
   "System_Byte" AT %MB0 : Byte;
END_VAR

VAR_GLOBAL CONSTANT   // PLC tag table "Tabella delle variabili standard"
   "CONST_dNumberOfHeadsCycle" : DInt := 7;   // Number of heads / Number of heads-1
   "CONST_dNumberOfHeads" : DInt := 8;   // Number of heads-1 / Number of heads
   "CONST_dPressureMax_MN" : DInt := 180000;   // Maximum allowable pressure [N/1000]
   "CONST_dPressureMin_MN" : DInt := 0;   // Minimum allowable pressure [N/1000]
   "CONST_dPressureMax_Unit" : DInt := 27648;   // Maximum allowable pressure Analog unit
   "CONST_dPressureMin_Unit" : DInt := 0;   // Minimum allowable pressure Analog unit
   "CONST_dFire_OnOff_MaxValue" : DInt := 5000;   // Fire ON OFF max value [mm/100]
   "CONST_dFire_OnOff_MinValue" : DInt := 0;   // Fire ON OFF min value [mm/100]
   "CONST_dPressureMax_Display_MN" : DInt := 180000;   // Maximum allowable pressure [N/1000]
   "CONST_dPressureMin_Display_MN" : DInt := 0;   // Minimum allowable pressure [N/1000]
   "CONST_dPressureMax_Display_Unit" : DInt := 27648;   // Maximum allowable pressure Analog unit
   "CONST_dPressureMin_Display_Unit" : DInt := 0;   // Minimum allowable pressure Analog unit
   "CONST_dPressureIncreasePneumatic_MN" : DInt := 250000;   // Pressure increse by cylinder [N/1000]
END_VAR

TYPE "ILx2T_Ref"
AUTHOR : SEMotion
FAMILY : LXM32
VERSION : 0.5
   STRUCT
      i_woDriveStatus : Word;
      i_by_ModeStatus : Byte;
      i_by_driveInput : Byte;
      i_wo_ActionWord : Word;
      i_wo_SpecialFunctions : Word;
      q_wo_dmControl : Word;
      q_dw_refA_16 : Word;
      q_dw_refB_32 : DWord;
      arOutputData : Array[0..7] of Byte;
      arInputData : Array[0..7] of Byte;
      stDriveStatus : Struct
         HaltActive : Bool;   // HALT is active
         reserved_Bit9 : Bool;
         reserved_Bit10 : Bool;
         reserved_Bit11 : Bool;
         reserved_Bit12 : Bool;
         x_Add : Bool;   // additional information
         x_End : Bool;   // OP mode finished - standstill
         x_Err : Bool;   // error
         state_Bit0 : Bool;   // Drive state bit 0
         state_Bit1 : Bool;   // Drive state bit 1
         state_Bit2 : Bool;   // Drive state bit 2
         state_Bit3 : Bool;   // Drive state bit 3
         reseverd_Bit4 : Bool;
         reserved_Bit5 : Bool;
         FaultActive : Bool;   // FAULT is active
         WarningActive : Bool;   // WARNING is active
      END_STRUCT;
      st_ModeStatus : Struct
         Mode_0 : Bool;   // Actual OP mode bit 0
         Mode_1 : Bool;   // Actual OP mode bit 1
         Mode_2 : Bool;   // Actual OP mode bit 2
         Mode_3 : Bool;   // Actual OP mode bit 3
         reserved : Bool;
         Reference_OK : Bool;   // drive is referenced
         ModeError : Bool;   // Status mode error
         ModeToggle : Bool;   // Status mode toggle
      END_STRUCT;
      st_ActionWord : Struct
         MotionNegative : Bool;   // negative direction
         InsidePosWindow : Bool;   // Inside Position Window
         reserved_Bit10 : Bool;
         TargetVelocityZero : Bool;   // Target velocity is zero
         Decelerating : Bool;
         Accelerating : Bool;
         ConstantVelocity : Bool;
         reserved_Bit15 : Bool;
         Reserved : Bool;
         Reserved_1 : Bool;
         Reserved_2 : Bool;
         Reserved_3 : Bool;
         Reserved_4 : Bool;
         Reserved_5 : Bool;
         MotionZero : Bool;   // Motion zero, actual velocity is zero
         MotionPositive : Bool;   // motor is moving in positiove direction
      END_STRUCT;
      st_SpecFunctions : Struct
         reserved_4 : Bool;   // Capture counter channel 1 bit 0
         reserved_5 : Bool;   // Capture counter channel 1 bit 1
         reserved_6 : Bool;   // Capture counter channel 2 bit 0
         reserved_7 : Bool;   // Capture counter channel 2 bit 1
         reserved_12 : Bool;
         reserved_13 : Bool;
         reserved_14 : Bool;
         reserved_15 : Bool;
         CAP1_0 : Bool;   // Actual OP mode bit 0
         CAP1_1 : Bool;   // Actual OP mode bit 1
         CAP2_0 : Bool;   // Actual OP mode bit 2
         CAP2_1 : Bool;   // Actual OP mode bit 3
         reserved : Bool;   // Actual OP mode bit 4
         reserved_1 : Bool;   // Status ModeDataError
         reserved_2 : Bool;   // Status mode error
         reserved_3 : Bool;   // Status mode toggle
      END_STRUCT;
      InitAccessID : Int;   // AccessID counter for INIT
      ProChAccessID : Int;   // Access ID Processchannel
      ParChAccessID : Int;   // Access ID Parameterchannel
      x_QuickStopInt : Bool;   // Library internal QuickStop Command
      x_FaultResetInt : Bool;   // Library internal FaultReset Command
      x_Set_HALT_Int : Bool;   // Library internal Set HALT Command
      x_Clear_HALT_Int : Bool;   // Library internal Clear HALT Command
      x_Continue_Int : Bool;   // Library internal HALT Contimue Command
      by_OP_ModeAct : Byte;   // Status - Actual operation mode
      x_IO_1 : Bool;   // Status of digital IO 1 (Bit 0)
      x_IO_2 : Bool;   // Status of digital IO 2 (Bit 1)
      x_IO_3 : Bool;   // Status of digital IO 3 (Bit 2)
      x_IO_4 : Bool;   // Status of digital IO 4 (Bit 3)
      x_STO_A : Bool;   // Status of Safe Torque Off Channel A
      x_STO_B : Bool;   // Status of Safe Torque Off Channel B
      x_reserved_6 : Bool;
      x_reserved_7 : Bool;
      x_CommandWriteParameter : Bool;
      x_CommandReadParameter : Bool;
      x_StatusReadParameter_OK : Bool;
      x_StatusReadParameter_Error : Bool;
      x_Status_WriteParameter_OK : Bool;
      x_Status_WriteParameter_Error : Bool;
      di_ParameterReadValue : DInt;
      di_ParameterWriteValue : DInt;
      udi_ModbusAddress_Read : UDInt;
      udi_ModbusAddress_Write : UDInt;
   END_STRUCT;
END_TYPE

TYPE "UDT_DataManager_HeadsBuffer"
VERSION : 0.1
   STRUCT
      rgdMissionID : Array[0..20] of DInt;   // Head#x mission ID
      rgdRequestPosition_cmm : Array[0..20] of DInt;   // Head#x request position [mm/100]
      rgdFireRequest : Array[0..20] of DInt;   // Head#x fire request
      dNumberOfElement : DInt;   // Number of element inside the buffer
   END_STRUCT;
END_TYPE

TYPE "UDT_DataManager_Insert"
VERSION : 0.1
   STRUCT
      dMissionCode : DInt;   // Mission code
      dMissionStart_cmm : DInt;   // Mission counter start [mm/100]
      dMissionEnd_cmm : DInt;   // Mission counter end [mm/100]
      rgxFireRequest : Array[0.."CONST_dNumberOfHeadsCycle"] of Bool;   // Fire request missions
      rgdHeadsPosition_cmm : Array[0.."CONST_dNumberOfHeadsCycle"] of DInt;   // Head#x position request [mm/100]
      xNewMission : Bool;   // New mission available
      xSystemReset : Bool;   // System reset
      rgdArmONReaction_ms : Array[0.."CONST_dNumberOfHeadsCycle"] of DInt;   // Head#x arm ON reaction [ms]
      rgdArmOFFReaction_ms : Array[0.."CONST_dNumberOfHeadsCycle"] of DInt;   // Head#x arm OFF reaction [ms]
      rgdFireONReaction_ms : Array[0.."CONST_dNumberOfHeadsCycle"] of DInt;   // Head#x fire ON reaction [ms]
      rgdFireOFFReaction_ms : Array[0.."CONST_dNumberOfHeadsCycle"] of DInt;   // Head#x fire OFF reaction [ms]
      rgdOilDelayStart_ms : Array[0.."CONST_dNumberOfHeadsCycle"] of DInt;   // Head#x oil delay start [ms]
      rgdOilDelayEnd_ms : Array[0.."CONST_dNumberOfHeadsCycle"] of DInt;   // Head#x oil advance end [ms]
      rgdFireONDelayStart_cmm : Array[0.."CONST_dNumberOfHeadsCycle"] of DInt;   // Head#x fire ON delay start [mm/100]
      rgdFireOFFDelayEnd_cmm : Array[0.."CONST_dNumberOfHeadsCycle"] of DInt;   // Head#x fire OFF delay end [mm/100]
   END_STRUCT;
END_TYPE

TYPE "UDT_DataManager"
VERSION : 0.1
   STRUCT
      tInputData : "UDT_DataManager_Insert";   // Manager input data
      tOutputData : "UDT_DataManager_Output";   // Manager output data
      dInterruptNumMissionTank : DInt;   // Number of mission fire inside the tank
      rgtInterruptMissionTank : Array[0..20] of "UDT_DataManager_Tank";   // Array of fire missions
      rgtOilList : Array[0.."CONST_dNumberOfHeadsCycle"] of "UDT_DataManager_HeadsBuffer";   // Oil list manager
      rgtArmList : Array[0.."CONST_dNumberOfHeadsCycle"] of "UDT_DataManager_HeadsBuffer";   // Arm list manager
   END_STRUCT;
END_TYPE

TYPE "UDT_DataManager_Output"